(* Logix 5000 project; controller FV vendor 1 type 14 code 217 rev 31.11; software revision 31.00; part 25 of 63 *)
(* tags used below, declared in another part *)
   CheckTimeMask : INT;
   Delphi_Does_Eng_Func : BOOL;
   FR_FV26_AV08 : PlantItem;   // FV26_AV08
   FR_FV27_AV08 : PlantItem;   // FV27_AV08
   FR_FV31_AV01 : PlantItem;   // FV31_AV01
   FR_FV31_AV04 : PlantItem;   // FV31_AV04
   FR_FV31_AV05 : PlantItem;   // FV31_AV05
   FR_FV31_AV06 : PlantItem;   // FV31_AV06
   FR_FV31_AV07 : PlantItem;   // FV31_AV07
   FR_N255 : INT[265];   // CHECKWORDS
   FR_VB3_AV01 : PlantItem;   // VB3_AV01
   FR_VB3_AV02 : PlantItem;   // VB3_AV02
   FR_VB3_AV03 : PlantItem;   // VB3_AV03
   FR_VB3_AV04 : PlantItem;   // VB3_AV04
   FR_VB3_AV05 : PlantItem;   // VB3_AV05
   FR_VB4_AV16 : PlantItem;   // VB4_AV16
   TempChecktime : DINT;
(* FR_Common, continued *)

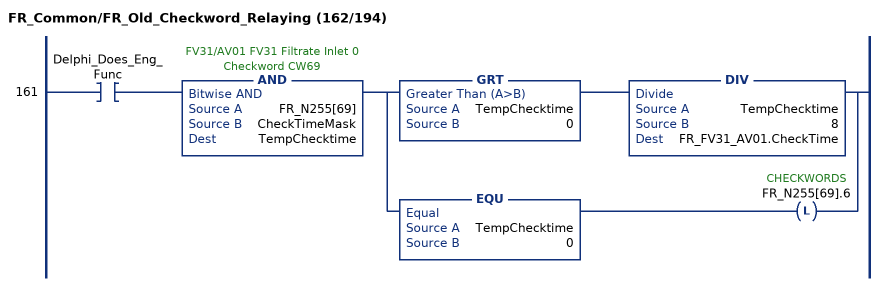
   [picture p466: FR_Common/FR_Old_Checkword_Relaying rungs 161-161]
   161: XIC(Delphi_Does_Eng_Func)AND(FR_N255[69],CheckTimeMask,TempChecktime)[GRT(TempChecktime,0) DIV(TempChecktime,8,FR_FV31_AV01.CheckTime) ,EQU(TempChecktime,0) OTL(FR_N255[69].6) ];
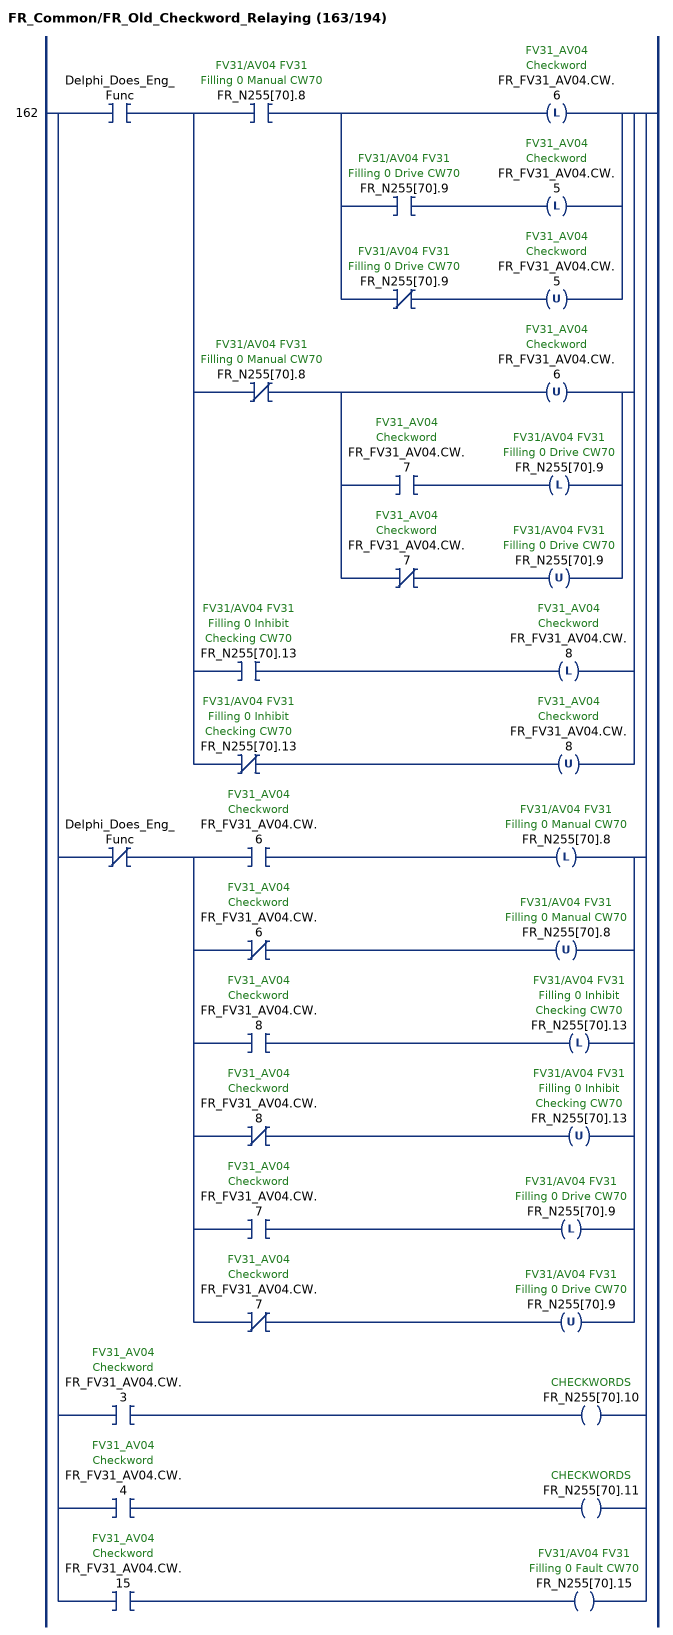
   162: [XIC(Delphi_Does_Eng_Func) [[XIC(FR_N255[70].8) [OTL(FR_FV31_AV04.CW.6) ,XIC(FR_N255[70].9) OTL(FR_FV31_AV04.CW.5) ,XIO(FR_N255[70].9) OTU(FR_FV31_AV04.CW.5) ] ,XIO(FR_N255[70].8) [OTU(FR_FV31_AV04.CW.6) ,[XIC(FR_FV31_AV04.CW.7) OTL(FR_N255[70].9) ,XIO(FR_FV31_AV04.CW.7) OTU(FR_N255[70].9) ] ] ] ,[XIC(FR_N255[70].13) OTL(FR_FV31_AV04.CW.8) ,XIO(FR_N255[70].13) OTU(FR_FV31_AV04.CW.8) ] ] ,XIO(Delphi_Does_Eng_Func) [[XIC(FR_FV31_AV04.CW.6) OTL(FR_N255[70].8) ,XIO(FR_FV31_AV04.CW.6) OTU(FR_N255[70].8) ] ,[XIC(FR_FV31_AV04.CW.8) OTL(FR_N255[70].13) ,XIO(FR_FV31_AV04.CW.8) OTU(FR_N255[70].13) ] ,[XIC(FR_FV31_AV04.CW.7) OTL(FR_N255[70].9) ,XIO(FR_FV31_AV04.CW.7) OTU(FR_N255[70].9) ] ] ,XIC(FR_FV31_AV04.CW.3) OTE(FR_N255[70].10) ,XIC(FR_FV31_AV04.CW.4) OTE(FR_N255[70].11) ,XIC(FR_FV31_AV04.CW.15) OTE(FR_N255[70].15) ];
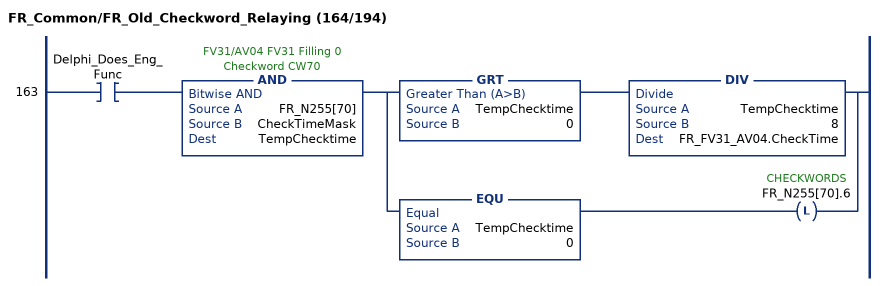
   163: XIC(Delphi_Does_Eng_Func)AND(FR_N255[70],CheckTimeMask,TempChecktime)[GRT(TempChecktime,0) DIV(TempChecktime,8,FR_FV31_AV04.CheckTime) ,EQU(TempChecktime,0) OTL(FR_N255[70].6) ];
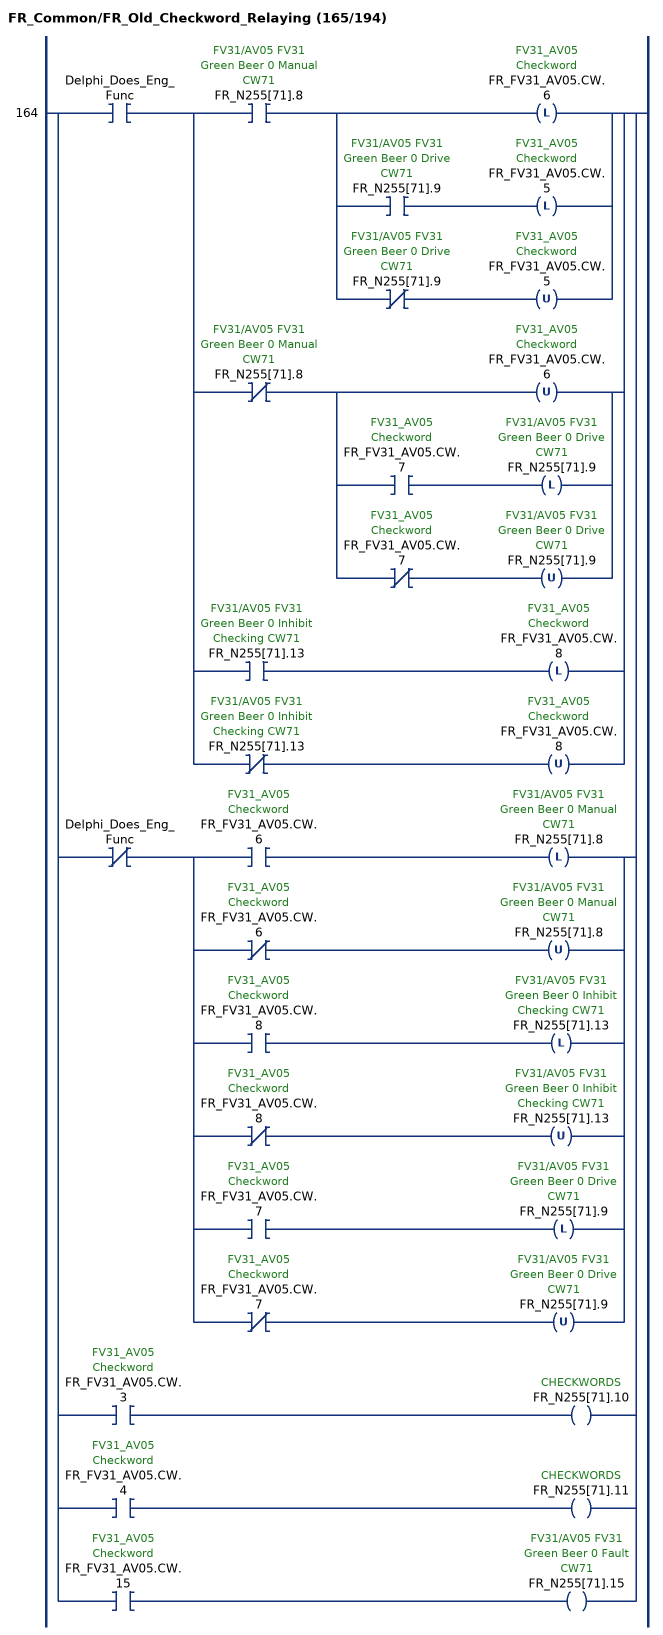
   164: [XIC(Delphi_Does_Eng_Func) [[XIC(FR_N255[71].8) [OTL(FR_FV31_AV05.CW.6) ,XIC(FR_N255[71].9) OTL(FR_FV31_AV05.CW.5) ,XIO(FR_N255[71].9) OTU(FR_FV31_AV05.CW.5) ] ,XIO(FR_N255[71].8) [OTU(FR_FV31_AV05.CW.6) ,[XIC(FR_FV31_AV05.CW.7) OTL(FR_N255[71].9) ,XIO(FR_FV31_AV05.CW.7) OTU(FR_N255[71].9) ] ] ] ,[XIC(FR_N255[71].13) OTL(FR_FV31_AV05.CW.8) ,XIO(FR_N255[71].13) OTU(FR_FV31_AV05.CW.8) ] ] ,XIO(Delphi_Does_Eng_Func) [[XIC(FR_FV31_AV05.CW.6) OTL(FR_N255[71].8) ,XIO(FR_FV31_AV05.CW.6) OTU(FR_N255[71].8) ] ,[XIC(FR_FV31_AV05.CW.8) OTL(FR_N255[71].13) ,XIO(FR_FV31_AV05.CW.8) OTU(FR_N255[71].13) ] ,[XIC(FR_FV31_AV05.CW.7) OTL(FR_N255[71].9) ,XIO(FR_FV31_AV05.CW.7) OTU(FR_N255[71].9) ] ] ,XIC(FR_FV31_AV05.CW.3) OTE(FR_N255[71].10) ,XIC(FR_FV31_AV05.CW.4) OTE(FR_N255[71].11) ,XIC(FR_FV31_AV05.CW.15) OTE(FR_N255[71].15) ];
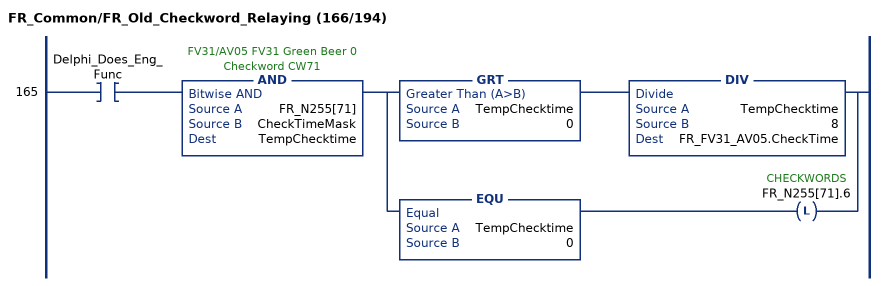
   165: XIC(Delphi_Does_Eng_Func)AND(FR_N255[71],CheckTimeMask,TempChecktime)[GRT(TempChecktime,0) DIV(TempChecktime,8,FR_FV31_AV05.CheckTime) ,EQU(TempChecktime,0) OTL(FR_N255[71].6) ];
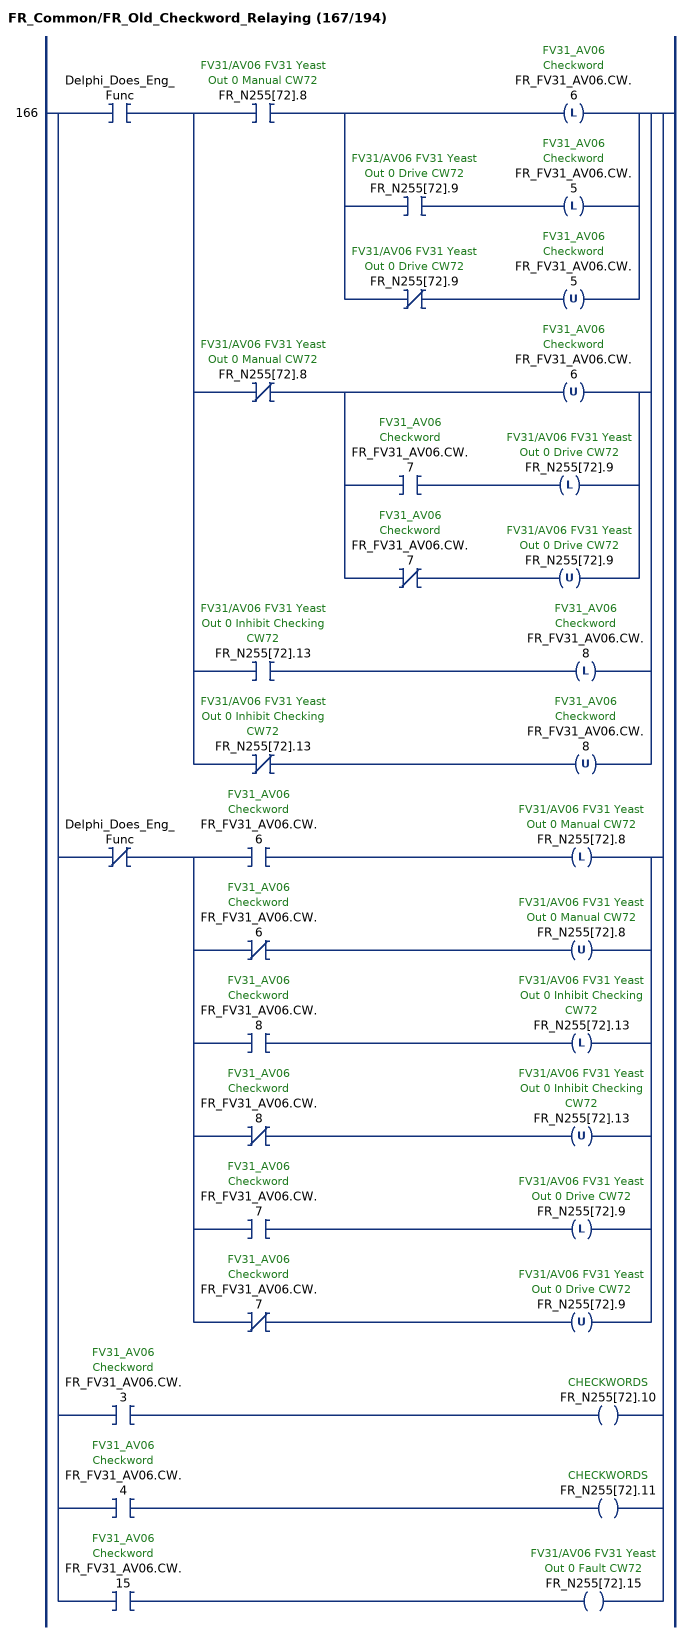
   166: [XIC(Delphi_Does_Eng_Func) [[XIC(FR_N255[72].8) [OTL(FR_FV31_AV06.CW.6) ,XIC(FR_N255[72].9) OTL(FR_FV31_AV06.CW.5) ,XIO(FR_N255[72].9) OTU(FR_FV31_AV06.CW.5) ] ,XIO(FR_N255[72].8) [OTU(FR_FV31_AV06.CW.6) ,[XIC(FR_FV31_AV06.CW.7) OTL(FR_N255[72].9) ,XIO(FR_FV31_AV06.CW.7) OTU(FR_N255[72].9) ] ] ] ,[XIC(FR_N255[72].13) OTL(FR_FV31_AV06.CW.8) ,XIO(FR_N255[72].13) OTU(FR_FV31_AV06.CW.8) ] ] ,XIO(Delphi_Does_Eng_Func) [[XIC(FR_FV31_AV06.CW.6) OTL(FR_N255[72].8) ,XIO(FR_FV31_AV06.CW.6) OTU(FR_N255[72].8) ] ,[XIC(FR_FV31_AV06.CW.8) OTL(FR_N255[72].13) ,XIO(FR_FV31_AV06.CW.8) OTU(FR_N255[72].13) ] ,[XIC(FR_FV31_AV06.CW.7) OTL(FR_N255[72].9) ,XIO(FR_FV31_AV06.CW.7) OTU(FR_N255[72].9) ] ] ,XIC(FR_FV31_AV06.CW.3) OTE(FR_N255[72].10) ,XIC(FR_FV31_AV06.CW.4) OTE(FR_N255[72].11) ,XIC(FR_FV31_AV06.CW.15) OTE(FR_N255[72].15) ];
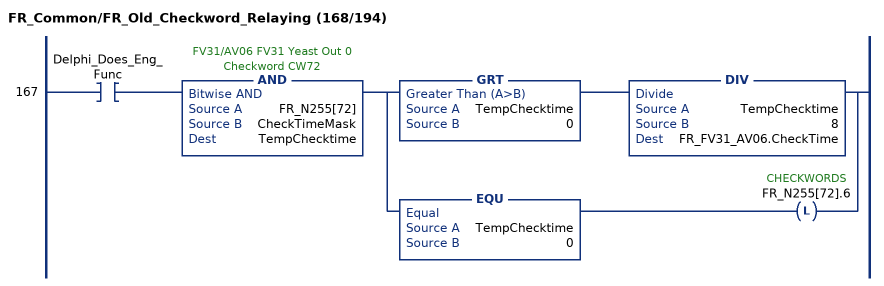
   167: XIC(Delphi_Does_Eng_Func)AND(FR_N255[72],CheckTimeMask,TempChecktime)[GRT(TempChecktime,0) DIV(TempChecktime,8,FR_FV31_AV06.CheckTime) ,EQU(TempChecktime,0) OTL(FR_N255[72].6) ];
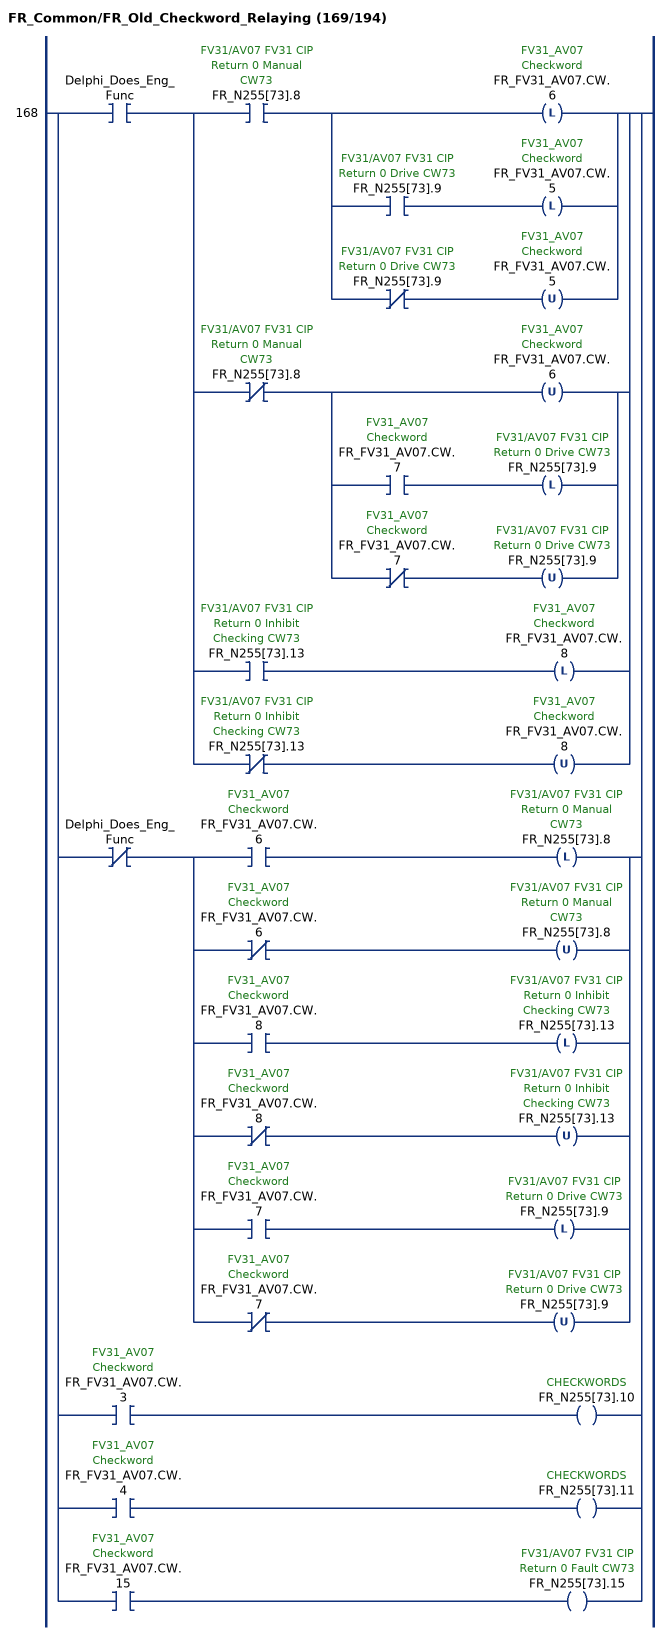
   168: [XIC(Delphi_Does_Eng_Func) [[XIC(FR_N255[73].8) [OTL(FR_FV31_AV07.CW.6) ,XIC(FR_N255[73].9) OTL(FR_FV31_AV07.CW.5) ,XIO(FR_N255[73].9) OTU(FR_FV31_AV07.CW.5) ] ,XIO(FR_N255[73].8) [OTU(FR_FV31_AV07.CW.6) ,[XIC(FR_FV31_AV07.CW.7) OTL(FR_N255[73].9) ,XIO(FR_FV31_AV07.CW.7) OTU(FR_N255[73].9) ] ] ] ,[XIC(FR_N255[73].13) OTL(FR_FV31_AV07.CW.8) ,XIO(FR_N255[73].13) OTU(FR_FV31_AV07.CW.8) ] ] ,XIO(Delphi_Does_Eng_Func) [[XIC(FR_FV31_AV07.CW.6) OTL(FR_N255[73].8) ,XIO(FR_FV31_AV07.CW.6) OTU(FR_N255[73].8) ] ,[XIC(FR_FV31_AV07.CW.8) OTL(FR_N255[73].13) ,XIO(FR_FV31_AV07.CW.8) OTU(FR_N255[73].13) ] ,[XIC(FR_FV31_AV07.CW.7) OTL(FR_N255[73].9) ,XIO(FR_FV31_AV07.CW.7) OTU(FR_N255[73].9) ] ] ,XIC(FR_FV31_AV07.CW.3) OTE(FR_N255[73].10) ,XIC(FR_FV31_AV07.CW.4) OTE(FR_N255[73].11) ,XIC(FR_FV31_AV07.CW.15) OTE(FR_N255[73].15) ];
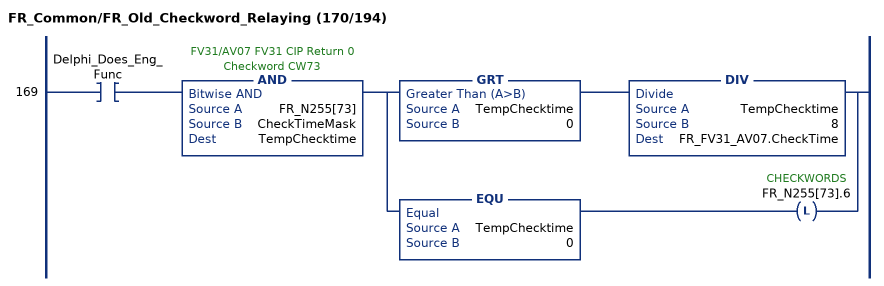
   169: XIC(Delphi_Does_Eng_Func)AND(FR_N255[73],CheckTimeMask,TempChecktime)[GRT(TempChecktime,0) DIV(TempChecktime,8,FR_FV31_AV07.CheckTime) ,EQU(TempChecktime,0) OTL(FR_N255[73].6) ];
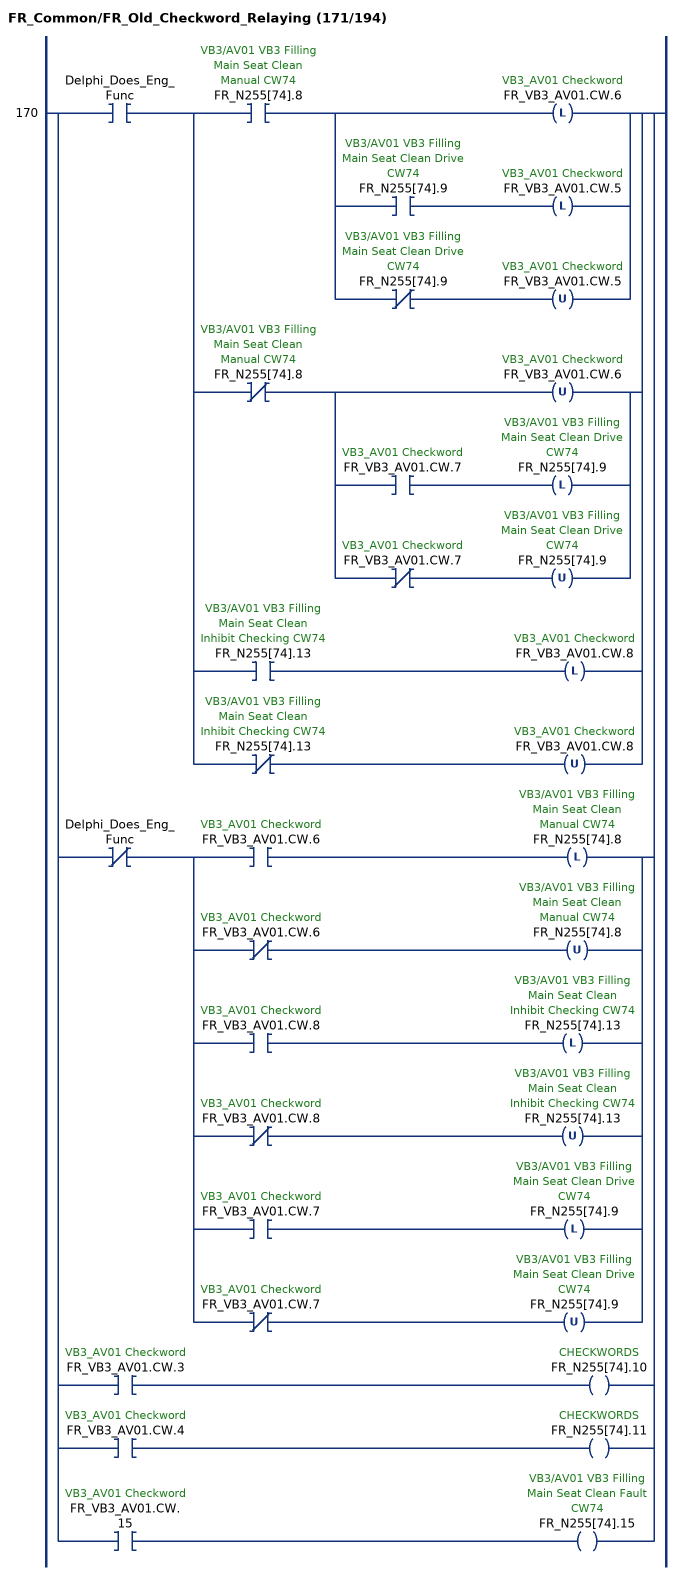
   170: [XIC(Delphi_Does_Eng_Func) [[XIC(FR_N255[74].8) [OTL(FR_VB3_AV01.CW.6) ,XIC(FR_N255[74].9) OTL(FR_VB3_AV01.CW.5) ,XIO(FR_N255[74].9) OTU(FR_VB3_AV01.CW.5) ] ,XIO(FR_N255[74].8) [OTU(FR_VB3_AV01.CW.6) ,[XIC(FR_VB3_AV01.CW.7) OTL(FR_N255[74].9) ,XIO(FR_VB3_AV01.CW.7) OTU(FR_N255[74].9) ] ] ] ,[XIC(FR_N255[74].13) OTL(FR_VB3_AV01.CW.8) ,XIO(FR_N255[74].13) OTU(FR_VB3_AV01.CW.8) ] ] ,XIO(Delphi_Does_Eng_Func) [[XIC(FR_VB3_AV01.CW.6) OTL(FR_N255[74].8) ,XIO(FR_VB3_AV01.CW.6) OTU(FR_N255[74].8) ] ,[XIC(FR_VB3_AV01.CW.8) OTL(FR_N255[74].13) ,XIO(FR_VB3_AV01.CW.8) OTU(FR_N255[74].13) ] ,[XIC(FR_VB3_AV01.CW.7) OTL(FR_N255[74].9) ,XIO(FR_VB3_AV01.CW.7) OTU(FR_N255[74].9) ] ] ,XIC(FR_VB3_AV01.CW.3) OTE(FR_N255[74].10) ,XIC(FR_VB3_AV01.CW.4) OTE(FR_N255[74].11) ,XIC(FR_VB3_AV01.CW.15) OTE(FR_N255[74].15) ];
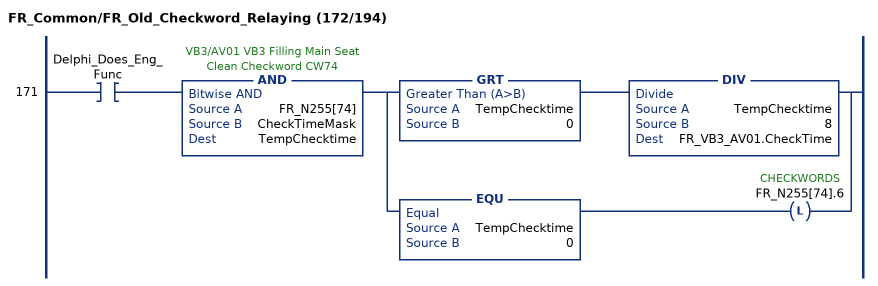
   171: XIC(Delphi_Does_Eng_Func)AND(FR_N255[74],CheckTimeMask,TempChecktime)[GRT(TempChecktime,0) DIV(TempChecktime,8,FR_VB3_AV01.CheckTime) ,EQU(TempChecktime,0) OTL(FR_N255[74].6) ];
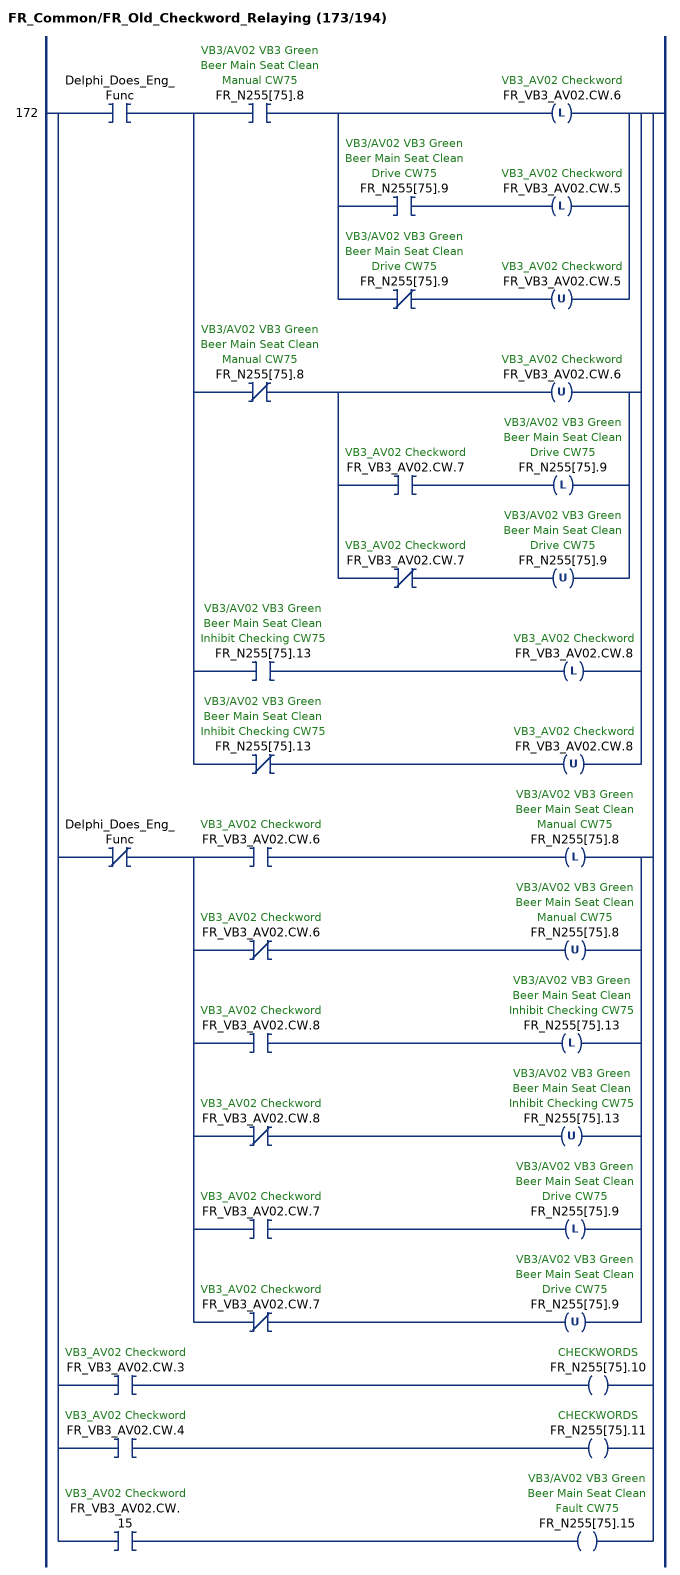
   172: [XIC(Delphi_Does_Eng_Func) [[XIC(FR_N255[75].8) [OTL(FR_VB3_AV02.CW.6) ,XIC(FR_N255[75].9) OTL(FR_VB3_AV02.CW.5) ,XIO(FR_N255[75].9) OTU(FR_VB3_AV02.CW.5) ] ,XIO(FR_N255[75].8) [OTU(FR_VB3_AV02.CW.6) ,[XIC(FR_VB3_AV02.CW.7) OTL(FR_N255[75].9) ,XIO(FR_VB3_AV02.CW.7) OTU(FR_N255[75].9) ] ] ] ,[XIC(FR_N255[75].13) OTL(FR_VB3_AV02.CW.8) ,XIO(FR_N255[75].13) OTU(FR_VB3_AV02.CW.8) ] ] ,XIO(Delphi_Does_Eng_Func) [[XIC(FR_VB3_AV02.CW.6) OTL(FR_N255[75].8) ,XIO(FR_VB3_AV02.CW.6) OTU(FR_N255[75].8) ] ,[XIC(FR_VB3_AV02.CW.8) OTL(FR_N255[75].13) ,XIO(FR_VB3_AV02.CW.8) OTU(FR_N255[75].13) ] ,[XIC(FR_VB3_AV02.CW.7) OTL(FR_N255[75].9) ,XIO(FR_VB3_AV02.CW.7) OTU(FR_N255[75].9) ] ] ,XIC(FR_VB3_AV02.CW.3) OTE(FR_N255[75].10) ,XIC(FR_VB3_AV02.CW.4) OTE(FR_N255[75].11) ,XIC(FR_VB3_AV02.CW.15) OTE(FR_N255[75].15) ];